// TIA Portal project "forward_reverse" (V16)

(* hardware
DEVICE "S7-1200 station_1"  S7-1200 Station
   slot 0: "Rack_0"  S7-1200 Rack  Rack  V1.0
   slot 1: "PLC_1"  CPU 1212C DC/DC/Rly  6ES7 212-1HE40-0XB0  V4.4
DEVICE "HMI_1"  TP700 Comfort
   slot 0: "HMI_1"  TP700 Comfort  6AV2 124-0GC01-0AX0  16.0.0.0
   slot 1: "HMI_RT_1"  TP700 Comfort  6AV2 124-0GC01-0AX0  16.0.0.0
   slot 5: "HMI_1.IE_CP_1"  PROFINET Interface  16.0.0.0
      slot 1: "PROFINET Interface_1"  PROFINET Interface
         slot 1: "Port_1"  Port
         slot 2: "Port_2"  Port
   slot 7: "HMI_1.MPI/DP_CP_1"  MPI/DP Interface  16.0.0.0
*)

// ===== PLC "PLC_1"  CPU 1212C DC/DC/Rly =====

VAR_GLOBAL   // PLC tag table "Default tag table"
   "PB_MOVE_R" AT %I0.0 : Bool;
   "PB_MOVE_F" AT %I0.1 : Bool;
   "PB_STOP" AT %I0.2 : Bool;
   "PB_EMERGENCY" AT %I0.3 : Bool;
   "PB_RESET" AT %I0.4 : Bool;
   "SENSOR_HOME" AT %I0.5 : Bool;
   "SENSOR_FINISH" AT %I0.6 : Bool;
   "COIL_R" AT %Q0.0 : Bool;
   "COIL_F" AT %Q0.1 : Bool;
   "COIL_EMERGENCY" AT %Q0.2 : Bool;
   "PB_RESET_COUNT" AT %I0.7 : Bool;
END_VAR

DATA_BLOCK "Inputs_DB"   // DB1
{ S7_Optimized_Access := 'FALSE' }
VERSION : 0.1
   VAR
      MOVE_R : Bool;
      MOVE_F : Bool;
      STOP : Bool;
      EMERGENCY : Bool;
      RESET : Bool;
      RESET_COUNT : Bool;
      SENSOR_HOME : Bool;
      SENSOR_FINISH : Bool;
   END_VAR
BEGIN
END_DATA_BLOCK

DATA_BLOCK "States_DB"   // DB2
{ S7_Optimized_Access := 'FALSE' }
VERSION : 0.1
   VAR
      COUNTING_READY : Bool;
      COUNTING_FINISHED : Bool;
      MOTOR_WIND_DOWN : Bool;
      EMERGENCY_STATE : Bool;
   END_VAR
BEGIN
END_DATA_BLOCK

DATA_BLOCK "CONVEYOR_OPERATION_DB"   // DB4
{ S7_Optimized_Access := 'TRUE' }
VERSION : 0.1
// stored: InstanceOfName CONVEYOR_OPERATION
"CONVEYOR_OPERATION"
BEGIN
END_DATA_BLOCK

DATA_BLOCK "HMI_DB"   // DB7
{ S7_Optimized_Access := 'FALSE' }
VERSION : 0.1
   VAR
      MOVE_FORWARD : Bool;
      MOVE_REVERSE : Bool;
      STOP : Bool;
      EMERGENCY : Bool;
      RESET : Bool;
      COUNT_VALUE : Int;
      RESET_COUNTER : Bool;
      COUNTING_FINISHED : Bool;
      FORWARD : Bool;
      REVERSE : Bool;
   END_VAR
BEGIN
END_DATA_BLOCK

// folder: System blocks/Program resources

DATA_BLOCK "COUNTING_PRODUCT_DB"   // DB3
{ S7_Optimized_Access := 'TRUE' }
AUTHOR : Simatic
FAMILY : IEC
NAME : CNTR
VERSION : 1.0
// stored: InstanceOfName IEC_COUNTER
"IEC_COUNTER"
BEGIN
   PV := 5;
END_DATA_BLOCK

DATA_BLOCK "WIND_DOWN_TIMER_DB"   // DB5
{ S7_Optimized_Access := 'TRUE' }
AUTHOR : Simatic
FAMILY : IEC
NAME : IEC_TMR
VERSION : 1.0
// stored: InstanceOfName IEC_TIMER
"IEC_TIMER"
BEGIN
   PT := T#5000ms;
END_DATA_BLOCK

DATA_BLOCK "REVERSE_TIMER_DB"   // DB6
{ S7_Optimized_Access := 'TRUE' }
AUTHOR : Simatic
FAMILY : IEC
NAME : IEC_TMR
VERSION : 1.0
// stored: InstanceOfName IEC_TIMER
"IEC_TIMER"
BEGIN
   PT := T#5000ms;
END_DATA_BLOCK

// folder: (top level)

FUNCTION_BLOCK "CONVEYOR_OPERATION"   // FB1, LAD
{ S7_Optimized_Access := 'TRUE' }
VERSION : 0.1
   VAR_INPUT
      EMERGENCY_STATE : Bool;
      MOTOR_WIND_DOWN : Bool;
      INTERLOCK_F : Bool;
      INTERLOCK_R : Bool;
      MOVE_F : Bool;
      MOVE_R : Bool;
      COIL_F : Bool;
   END_VAR
   VAR_OUTPUT
      COIL_F_OUT : Bool;
      COIL_F_HMI : Bool;
      COIL_R_OUT : Bool;
      COIL_R_HMI : Bool;
   END_VAR
BEGIN

REGION Network 1
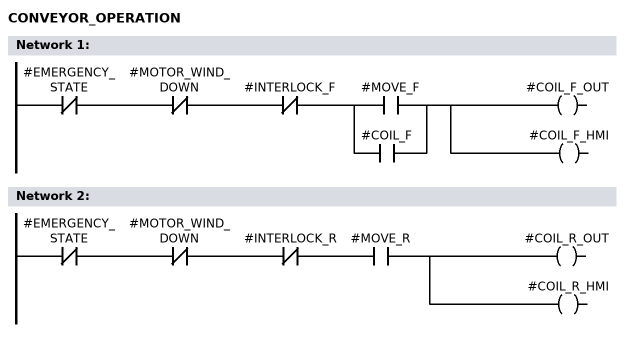
   RUNG wire#powerrail
      I_Contact( #EMERGENCY_STATE )
      I_Contact( #MOTOR_WIND_DOWN )
      I_Contact( #INTERLOCK_F )
      wire#w1
      Contact( #MOVE_F )
      wire#w2
      Coil( #COIL_F_OUT )
   END_RUNG
   RUNG wire#w1
      Contact( #COIL_F )
   END_RUNG wire#w2
   RUNG wire#w2
      Coil( #COIL_F_HMI )
   END_RUNG
   // the same network as SCL:
   #COIL_F_OUT := NOT #EMERGENCY_STATE AND NOT #MOTOR_WIND_DOWN AND NOT #INTERLOCK_F AND (#MOVE_F OR #COIL_F);
   #COIL_F_HMI := #COIL_F_OUT;
END_REGION

REGION Network 2
   RUNG wire#powerrail
      I_Contact( #EMERGENCY_STATE )
      I_Contact( #MOTOR_WIND_DOWN )
      I_Contact( #INTERLOCK_R )
      Contact( #MOVE_R )
      wire#w1
      Coil( #COIL_R_OUT )
   END_RUNG
   RUNG wire#w1
      Coil( #COIL_R_HMI )
   END_RUNG
   // the same network as SCL:
   #COIL_R_OUT := NOT #EMERGENCY_STATE AND NOT #MOTOR_WIND_DOWN AND NOT #INTERLOCK_R AND #MOVE_R;
   #COIL_R_HMI := #COIL_R_OUT;
END_REGION
END_FUNCTION_BLOCK

FUNCTION "I/O" : Void   // FC1, LAD
{ S7_Optimized_Access := 'TRUE' }
VERSION : 0.1
BEGIN

REGION Network 1
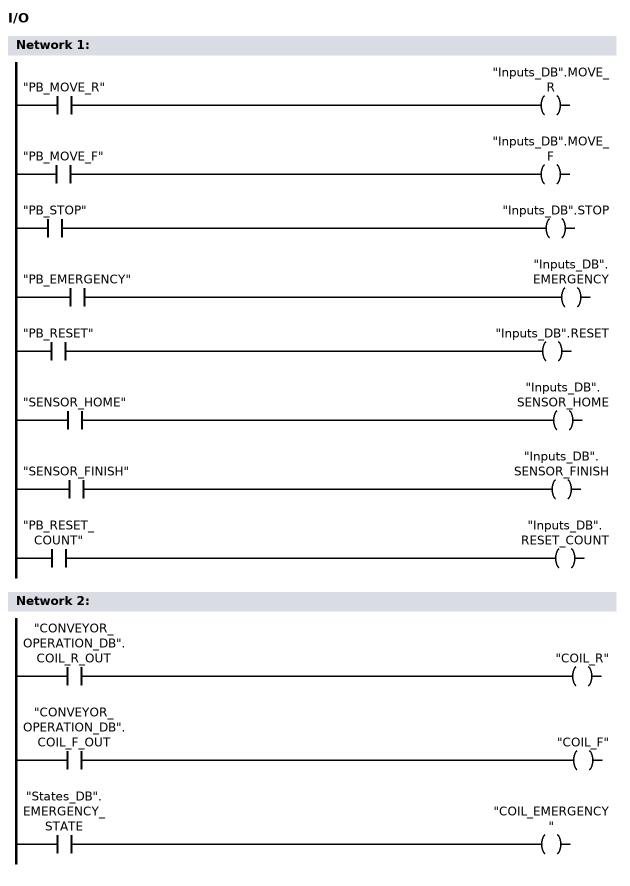
   RUNG wire#powerrail
      Contact( "PB_MOVE_R" )
      Coil( "Inputs_DB".MOVE_R )
   END_RUNG
   RUNG wire#powerrail
      Contact( "PB_MOVE_F" )
      Coil( "Inputs_DB".MOVE_F )
   END_RUNG
   RUNG wire#powerrail
      Contact( "PB_STOP" )
      Coil( "Inputs_DB".STOP )
   END_RUNG
   RUNG wire#powerrail
      Contact( "PB_EMERGENCY" )
      Coil( "Inputs_DB".EMERGENCY )
   END_RUNG
   RUNG wire#powerrail
      Contact( "PB_RESET" )
      Coil( "Inputs_DB".RESET )
   END_RUNG
   RUNG wire#powerrail
      Contact( "SENSOR_HOME" )
      Coil( "Inputs_DB".SENSOR_HOME )
   END_RUNG
   RUNG wire#powerrail
      Contact( "SENSOR_FINISH" )
      Coil( "Inputs_DB".SENSOR_FINISH )
   END_RUNG
   RUNG wire#powerrail
      Contact( "PB_RESET_COUNT" )
      Coil( "Inputs_DB".RESET_COUNT )
   END_RUNG
   // the same network as SCL:
   "Inputs_DB".MOVE_R := "PB_MOVE_R";
   "Inputs_DB".MOVE_F := "PB_MOVE_F";
   "Inputs_DB".STOP := "PB_STOP";
   "Inputs_DB".EMERGENCY := "PB_EMERGENCY";
   "Inputs_DB".RESET := "PB_RESET";
   "Inputs_DB".SENSOR_HOME := "SENSOR_HOME";
   "Inputs_DB".SENSOR_FINISH := "SENSOR_FINISH";
   "Inputs_DB".RESET_COUNT := "PB_RESET_COUNT";
END_REGION

REGION Network 2
   RUNG wire#powerrail
      Contact( "CONVEYOR_OPERATION_DB".COIL_R_OUT )
      Coil( "COIL_R" )
   END_RUNG
   RUNG wire#powerrail
      Contact( "CONVEYOR_OPERATION_DB".COIL_F_OUT )
      Coil( "COIL_F" )
   END_RUNG
   RUNG wire#powerrail
      Contact( "States_DB".EMERGENCY_STATE )
      Coil( "COIL_EMERGENCY" )
   END_RUNG
   // the same network as SCL:
   "COIL_R" := "CONVEYOR_OPERATION_DB".COIL_R_OUT;
   "COIL_F" := "CONVEYOR_OPERATION_DB".COIL_F_OUT;
   "COIL_EMERGENCY" := "States_DB".EMERGENCY_STATE;
END_REGION
END_FUNCTION

FUNCTION "COUNTING" : Void   // FC2, LAD
{ S7_Optimized_Access := 'TRUE' }
VERSION : 0.1
BEGIN

REGION Network 1
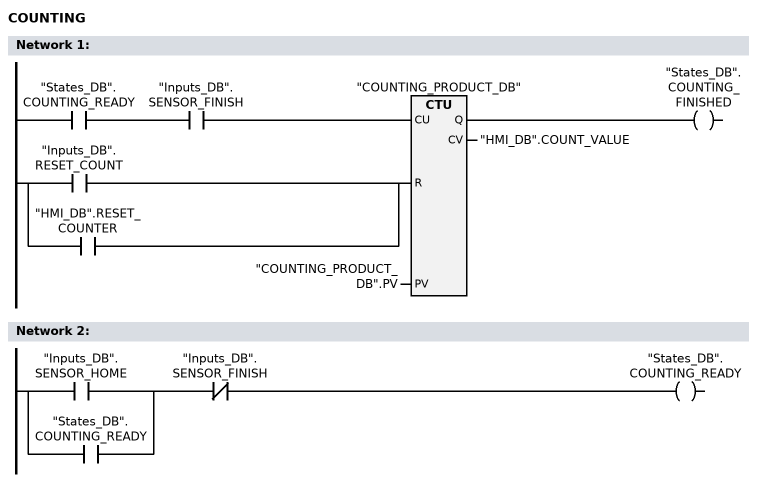
   "COUNTING_PRODUCT_DB".CTU(CU := "States_DB".COUNTING_READY AND "Inputs_DB".SENSOR_FINISH,
                           R := "Inputs_DB".RESET_COUNT OR "HMI_DB".RESET_COUNTER,
                           PV := "COUNTING_PRODUCT_DB".PV,
                           CV => "HMI_DB".COUNT_VALUE);
   "States_DB".COUNTING_FINISHED := "COUNTING_PRODUCT_DB".Q;
END_REGION

REGION Network 2
   RUNG wire#powerrail
      Contact( "Inputs_DB".SENSOR_HOME )
      wire#w1
      I_Contact( "Inputs_DB".SENSOR_FINISH )
      Coil( "States_DB".COUNTING_READY )
   END_RUNG
   RUNG wire#powerrail
      Contact( "States_DB".COUNTING_READY )
   END_RUNG wire#w1
   // the same network as SCL:
   "States_DB".COUNTING_READY := ("Inputs_DB".SENSOR_HOME OR "States_DB".COUNTING_READY) AND NOT "Inputs_DB".SENSOR_FINISH;
END_REGION
END_FUNCTION

FUNCTION "MOTOR_WIND_DOWN" : Void   // FC3, LAD
{ S7_Optimized_Access := 'TRUE' }
VERSION : 0.1
BEGIN

REGION Network 1
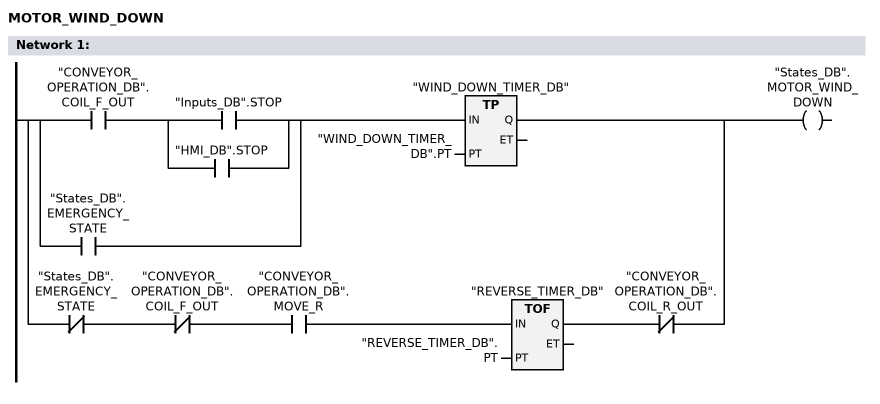
   "WIND_DOWN_TIMER_DB".TP(IN := ("CONVEYOR_OPERATION_DB".COIL_F_OUT AND ("Inputs_DB".STOP OR "HMI_DB".STOP)) OR "States_DB".EMERGENCY_STATE,
                           PT := "WIND_DOWN_TIMER_DB".PT);
   "REVERSE_TIMER_DB".TOF(IN := NOT "States_DB".EMERGENCY_STATE AND NOT "CONVEYOR_OPERATION_DB".COIL_F_OUT AND "CONVEYOR_OPERATION_DB".MOVE_R,
                          PT := "REVERSE_TIMER_DB".PT);
   "States_DB".MOTOR_WIND_DOWN := "WIND_DOWN_TIMER_DB".Q OR ("REVERSE_TIMER_DB".Q AND NOT "CONVEYOR_OPERATION_DB".COIL_R_OUT);
END_REGION
END_FUNCTION

ORGANIZATION_BLOCK "Main"   // OB1, LAD, ProgramCycle
TITLE = "Main Program Sweep (Cycle)"
{ S7_Optimized_Access := 'TRUE' }
VERSION : 0.1
   VAR_INPUT
      Initial_Call : Bool;   // Initial call of this OB
      Remanence : Bool;   // =True, if remanent data are available
   END_VAR
BEGIN

REGION Network 1
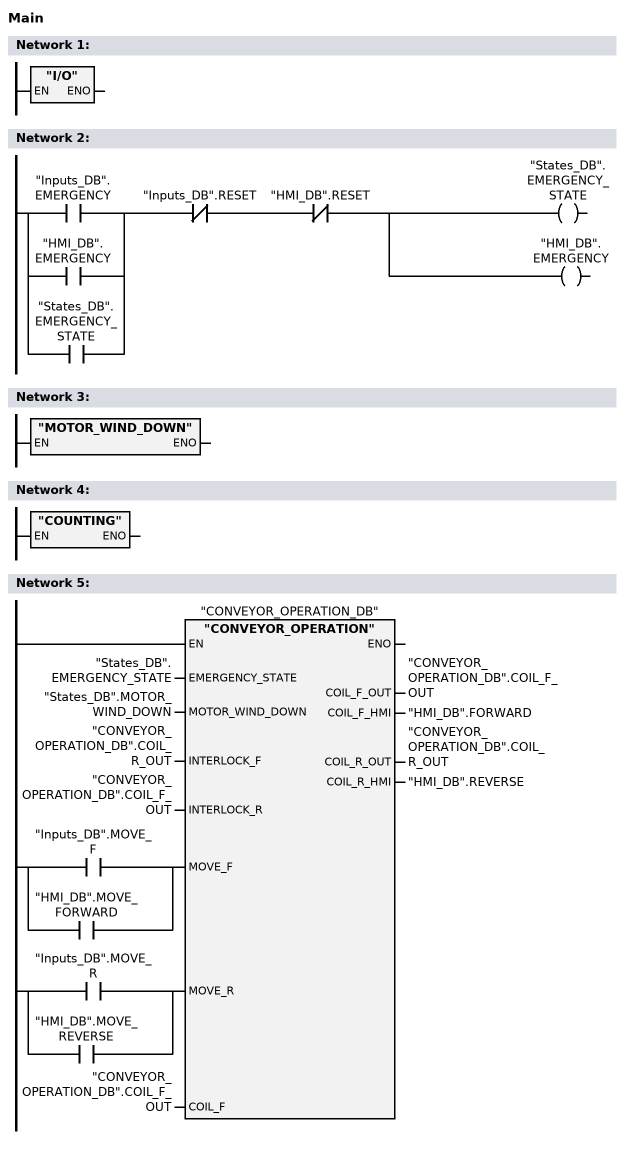
   RUNG wire#powerrail
      "I/O"()
   END_RUNG
   // the same network as SCL:
   "I/O"();
END_REGION

REGION Network 2
   RUNG wire#powerrail
      Contact( "Inputs_DB".EMERGENCY )
      wire#w1
      I_Contact( "Inputs_DB".RESET )
      I_Contact( "HMI_DB".RESET )
      wire#w2
      Coil( "States_DB".EMERGENCY_STATE )
   END_RUNG
   RUNG wire#powerrail
      Contact( "HMI_DB".EMERGENCY )
   END_RUNG wire#w1
   RUNG wire#powerrail
      Contact( "States_DB".EMERGENCY_STATE )
   END_RUNG wire#w1
   RUNG wire#w2
      Coil( "HMI_DB".EMERGENCY )
   END_RUNG
   // the same network as SCL:
   "States_DB".EMERGENCY_STATE := ("Inputs_DB".EMERGENCY OR "HMI_DB".EMERGENCY OR "States_DB".EMERGENCY_STATE) AND NOT "Inputs_DB".RESET AND NOT "HMI_DB".RESET;
   "HMI_DB".EMERGENCY := "States_DB".EMERGENCY_STATE;
END_REGION

REGION Network 3
   RUNG wire#powerrail
      "MOTOR_WIND_DOWN"()
   END_RUNG
   // the same network as SCL:
   "MOTOR_WIND_DOWN"();
END_REGION

REGION Network 4
   RUNG wire#powerrail
      "COUNTING"()
   END_RUNG
   // the same network as SCL:
   "COUNTING"();
END_REGION

REGION Network 5
   RUNG wire#powerrail
      "CONVEYOR_OPERATION_DB"(MOVE_F := wire#w1, MOVE_R := wire#w2, EMERGENCY_STATE := "States_DB".EMERGENCY_STATE, MOTOR_WIND_DOWN := "States_DB".MOTOR_WIND_DOWN, INTERLOCK_F := "CONVEYOR_OPERATION_DB".COIL_R_OUT, INTERLOCK_R := "CONVEYOR_OPERATION_DB".COIL_F_OUT, COIL_F := "CONVEYOR_OPERATION_DB".COIL_F_OUT, COIL_F_OUT => "CONVEYOR_OPERATION_DB".COIL_F_OUT, COIL_F_HMI => "HMI_DB".FORWARD, COIL_R_OUT => "CONVEYOR_OPERATION_DB".COIL_R_OUT, COIL_R_HMI => "HMI_DB".REVERSE)
   END_RUNG
   RUNG wire#powerrail
      Contact( "Inputs_DB".MOVE_F )
   END_RUNG wire#w1
   RUNG wire#powerrail
      Contact( "HMI_DB".MOVE_FORWARD )
   END_RUNG wire#w1
   RUNG wire#powerrail
      Contact( "Inputs_DB".MOVE_R )
   END_RUNG wire#w2
   RUNG wire#powerrail
      Contact( "HMI_DB".MOVE_REVERSE )
   END_RUNG wire#w2
   // the same network as SCL:
   "CONVEYOR_OPERATION_DB"(EMERGENCY_STATE := "States_DB".EMERGENCY_STATE,   // "CONVEYOR_OPERATION"
                           MOTOR_WIND_DOWN := "States_DB".MOTOR_WIND_DOWN,
                           INTERLOCK_F := "CONVEYOR_OPERATION_DB".COIL_R_OUT,
                           INTERLOCK_R := "CONVEYOR_OPERATION_DB".COIL_F_OUT,
                           MOVE_F := "Inputs_DB".MOVE_F OR "HMI_DB".MOVE_FORWARD,
                           MOVE_R := "Inputs_DB".MOVE_R OR "HMI_DB".MOVE_REVERSE,
                           COIL_F := "CONVEYOR_OPERATION_DB".COIL_F_OUT,
                           COIL_F_OUT => "CONVEYOR_OPERATION_DB".COIL_F_OUT,
                           COIL_F_HMI => "HMI_DB".FORWARD,
                           COIL_R_OUT => "CONVEYOR_OPERATION_DB".COIL_R_OUT,
                           COIL_R_HMI => "HMI_DB".REVERSE);
END_REGION
END_ORGANIZATION_BLOCK

(* ===== HMI "HMI_RT_1" =====
system functions are stored by id; their names below are inferred from use
connection "HMI_Connection_1": ETHERNET, S7_1200_OMS

HMI tags "Default tag table"
   "Tag_ScreenNumber" : UInt, internal
   "CONVEYOR_OPERATION_DB_COIL_F_OUT" : Bool = PLC CONVEYOR_OPERATION_DB.COIL_F_OUT, 1 s
   "CONVEYOR_OPERATION_DB_COIL_R_OUT" : Bool = PLC CONVEYOR_OPERATION_DB.COIL_R_OUT, 1 s
   "Inputs_DB_MOVE_F" : Bool = PLC Inputs_DB.MOVE_F AT %DB1.DBX0.1, 1 s
   "HMI_DB_REVERSE" : Bool = PLC HMI_DB.REVERSE AT %DB7.DBX4.3, 1 s
   "HMI_DB_FORWARD" : Bool = PLC HMI_DB.FORWARD AT %DB7.DBX4.2, 1 s
   "HMI_DB_MOVE_REVERSE" : Bool = PLC HMI_DB.MOVE_REVERSE AT %DB7.DBX0.1, 1 s
   "HMI_DB_MOVE_FORWARD" : Bool = PLC HMI_DB.MOVE_FORWARD AT %DB7.DBX0.0, 1 s
   "HMI_DB_STOP" : Bool = PLC HMI_DB.STOP AT %DB7.DBX0.2, 1 s
   "HMI_DB_EMERGENCY" : Bool = PLC HMI_DB.EMERGENCY AT %DB7.DBX0.3, 1 s
   "HMI_DB_RESET" : Bool = PLC HMI_DB.RESET AT %DB7.DBX0.4, 1 s
   "COUNTING_PRODUCT_DB_PV" : Int = PLC COUNTING_PRODUCT_DB.PV, 1 s
   "HMI_DB_COUNT_VALUE" : Int = PLC HMI_DB.COUNT_VALUE AT %DB7.DBW2, 1 s
   "COUNTING_PRODUCT_DB_CV" : Int = PLC COUNTING_PRODUCT_DB.CV, 1 s
   "HMI_DB_RESET_COUNTER" : Bool = PLC HMI_DB.RESET_COUNTER AT %DB7.DBX4.0, 1 s
   "States_DB_COUNTING_FINISHED" : Bool = PLC States_DB.COUNTING_FINISHED AT %DB2.DBX0.1, 1 s
   "States_DB_MOTOR_WIND_DOWN" : Bool = PLC States_DB.MOTOR_WIND_DOWN AT %DB2.DBX0.2, 1 s

screen "Root screen" 800x420, template "Template_1"
   on GenerateScreen: SetTag("Tag_ScreenNumber", 1)
   Circle "Circle_1" at 325,92 size 48x48
      Appearance <- "HMI_DB_REVERSE"
   Button "Button_1" at 513,218 size 96x32; TextOff 'FORWARD'
      on Press: function_b14e0dd5("HMI_DB_MOVE_FORWARD", 0)
   Button "Button_2" at 213,218 size 96x32; TextOff 'REVERSE'
      on Press: function_b14e0dd5("HMI_DB_MOVE_REVERSE", 0)
   Button "Button_3" at 364,218 size 96x32; TextOff 'STOP'
      on Press: function_b14e0dd5("HMI_DB_STOP", 0)
   Circle "Circle_2" at 453,92 size 48x48
      Appearance <- "HMI_DB_FORWARD"
   Circle "Circle_3" at 10,8 size 48x48
      Appearance <- "HMI_DB_EMERGENCY"
   Button "Button_4" at 10,67 size 129x32; TextOff 'EMERGENCY'
      on Press: function_b14e0dd5("HMI_DB_EMERGENCY", 0)
   Button "Button_5" at 10,129 size 96x32; TextOff 'RESET'
      on Press: function_b14e0dd5("HMI_DB_RESET", 0)
   Button "Button_6" at 609,27 size 163x40; TextOff 'COUNTER SCREEN'
      on Click: ActivateScreen("COUNTER SCREEN", 0)
   TextField "Text field_1" at 10,305 size 139x23; Text 'MOTOR READY'
   Rectangle "Rectangle_1" at 149,291 size 96x48
      Appearance <- "States_DB_MOTOR_WIND_DOWN"

Template "Template_1" 800x420
   Button "Exit" at 720,360 size 78x58; TextOff 'Exit'; PictureOff "ExitRuntime_TP700_Comfort_TR"; PictureOn "ExitRuntime_TP700_Comfort_TR"
      on Release: StopRuntime(0)
   Button "Template_Button" at 640,360 size 78x58; TextOff 'Text'
   Button "Template_Button_1" at 560,360 size 78x58; TextOff 'Text'
   Button "Template_Button_2" at 480,360 size 78x58; TextOff 'Text'
   Button "Template_Button_3" at 400,360 size 78x58; TextOff 'Text'
   Button "Template_Button_4" at 321,360 size 78x58; TextOff 'Text'
   Button "Template_Button_5" at 241,360 size 78x58; TextOff 'Text'
   Button "Template_Button_6" at 161,360 size 78x58; TextOff 'Text'
   Button "Alarms" at 81,360 size 78x58; TextOff 'Alarms'; PictureOff "AlarmDisplay_TP700_Comfort_TR"; PictureOn "AlarmDisplay_TP700_Comfort_TR"
      on Release: function_ef3f5d25("Alarm window_Unacknowledged", -1)
   Button "Start screen" at 1,360 size 78x58; TextOff 'Start screen'; PictureOff "NavigateHome_TP700_Comfort_TR"; PictureOn "NavigateHome_TP700_Comfort_TR"
      on Release: ActivateScreen("Root screen", 0)

screen "COUNTER SCREEN" 800x420
   Button "Button_1" at 667,33 size 96x32; TextOff 'HOME'
      on Click: ActivateScreen("Root screen", 0)
   TextField "Text field_1" at 69,135 size 132x23; Text 'SET COUNTER'
   TextField "Text field_2" at 69,175 size 157x23; Text 'COUNTER VALUE'
   IOField "I/O field_1" at 256,126 size 96x32; FormatPattern s99999
      ProcessValue <- "COUNTING_PRODUCT_DB_PV"
   IOField "I/O field_2" at 256,175 size 96x32; FormatPattern s99999
      ProcessValue <- "COUNTING_PRODUCT_DB_CV"
   Button "Button_2" at 125,230 size 181x32; TextOff 'RESET COUNTER'
      on Press: function_b14e0dd5("HMI_DB_RESET_COUNTER", 0)
   Circle "Circle_1" at 178,50 size 48x48
      Appearance <- "States_DB_COUNTING_FINISHED"
*)